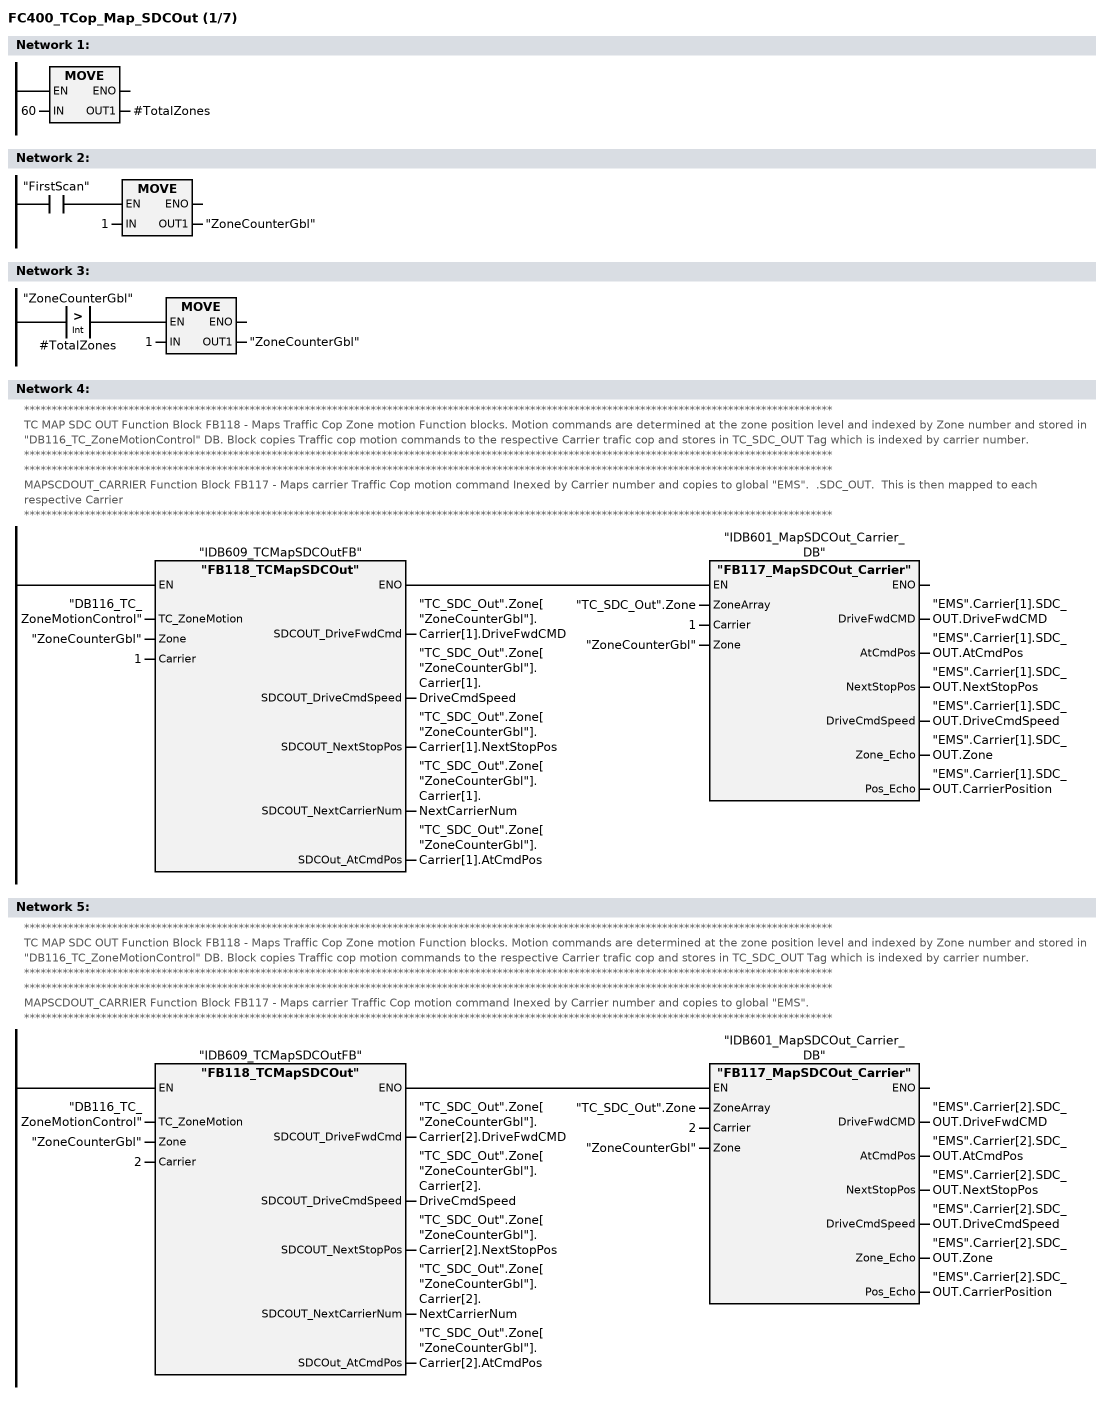
   RUNG wire#powerrail
      Move(in := 60, out1 => #TotalZones)
   END_RUNG
   // the same network as SCL:
   #TotalZones := 60;
END_REGION

REGION Network 2
   RUNG wire#powerrail
      Contact( "FirstScan" )
      Move(in := 1, out1 => "ZoneCounterGbl")
   END_RUNG
   // the same network as SCL:
   IF "FirstScan" THEN "ZoneCounterGbl" := 1; END_IF;
END_REGION

REGION Network 3
   RUNG wire#powerrail
      { S7_Templates := "SrcType := Int" } GT_Contact(in1 := "ZoneCounterGbl", in2 := #TotalZones)
      Move(in := 1, out1 => "ZoneCounterGbl")
   END_RUNG
   // the same network as SCL:
   IF "ZoneCounterGbl" > #TotalZones THEN "ZoneCounterGbl" := 1; END_IF;
END_REGION

REGION Network 4
   // ***************************************************************************************************************************************************
   // 
   // TC MAP SDC OUT Function Block FB118 - Maps Traffic Cop Zone motion Function blocks. Motion commands are determined at the zone position level and indexed by Zone number and stored in 
   //  "DB116_TC_ZoneMotionControl" DB. Block copies Traffic cop motion commands to the respective Carrier trafic cop and stores in TC_SDC_OUT Tag which is indexed by carrier number. 
   // 
   // ***************************************************************************************************************************************************
   // 
   // ***************************************************************************************************************************************************
   // 
   // MAPSCDOUT_CARRIER Function Block FB117 - Maps carrier Traffic Cop motion command Inexed by Carrier number and copies to global "EMS".  .SDC_OUT.  This is then mapped to each respective Carrier
   // 
   // ***************************************************************************************************************************************************
   RUNG wire#powerrail
      "IDB609_TCMapSDCOutFB"(TC_ZoneMotion := "DB116_TC_ZoneMotionControl", Zone := "ZoneCounterGbl", Carrier := 1, SDCOUT_DriveFwdCmd => "TC_SDC_Out".Zone["ZoneCounterGbl"].Carrier[1].DriveFwdCMD, SDCOUT_DriveCmdSpeed => "TC_SDC_Out".Zone["ZoneCounterGbl"].Carrier[1].DriveCmdSpeed, SDCOUT_NextStopPos => "TC_SDC_Out".Zone["ZoneCounterGbl"].Carrier[1].NextStopPos, SDCOUT_NextCarrierNum => "TC_SDC_Out".Zone["ZoneCounterGbl"].Carrier[1].NextCarrierNum, SDCOut_AtCmdPos => "TC_SDC_Out".Zone["ZoneCounterGbl"].Carrier[1].AtCmdPos)
      "IDB601_MapSDCOut_Carrier_DB"(ZoneArray := "TC_SDC_Out".Zone, Carrier := 1, Zone := "ZoneCounterGbl", DriveFwdCMD => "EMS".Carrier[1].SDC_OUT.DriveFwdCMD, AtCmdPos => "EMS".Carrier[1].SDC_OUT.AtCmdPos, NextStopPos => "EMS".Carrier[1].SDC_OUT.NextStopPos, DriveCmdSpeed => "EMS".Carrier[1].SDC_OUT.DriveCmdSpeed, Zone_Echo => "EMS".Carrier[1].SDC_OUT.Zone, Pos_Echo => "EMS".Carrier[1].SDC_OUT.CarrierPosition)
   END_RUNG
   // the same network as SCL:
   "IDB609_TCMapSDCOutFB"(TC_ZoneMotion := "DB116_TC_ZoneMotionControl",   // "FB118_TCMapSDCOut"
                          Zone := "ZoneCounterGbl",
                          Carrier := 1,
                          SDCOUT_DriveFwdCmd => "TC_SDC_Out".Zone["ZoneCounterGbl"].Carrier[1].DriveFwdCMD,
                          SDCOUT_DriveCmdSpeed => "TC_SDC_Out".Zone["ZoneCounterGbl"].Carrier[1].DriveCmdSpeed,
                          SDCOUT_NextStopPos => "TC_SDC_Out".Zone["ZoneCounterGbl"].Carrier[1].NextStopPos,
                          SDCOUT_NextCarrierNum => "TC_SDC_Out".Zone["ZoneCounterGbl"].Carrier[1].NextCarrierNum,
                          SDCOut_AtCmdPos => "TC_SDC_Out".Zone["ZoneCounterGbl"].Carrier[1].AtCmdPos,
                          ENO => #_w1);
   IF #_w1 THEN
       "IDB601_MapSDCOut_Carrier_DB"(ZoneArray := "TC_SDC_Out".Zone,   // "FB117_MapSDCOut_Carrier"
                               Carrier := 1,
                               Zone := "ZoneCounterGbl",
                               DriveFwdCMD => "EMS".Carrier[1].SDC_OUT.DriveFwdCMD,
                               AtCmdPos => "EMS".Carrier[1].SDC_OUT.AtCmdPos,
                               NextStopPos => "EMS".Carrier[1].SDC_OUT.NextStopPos,
                               DriveCmdSpeed => "EMS".Carrier[1].SDC_OUT.DriveCmdSpeed,
                               Zone_Echo => "EMS".Carrier[1].SDC_OUT.Zone,
                               Pos_Echo => "EMS".Carrier[1].SDC_OUT.CarrierPosition);
   END_IF;
END_REGION

REGION Network 5
   // ***************************************************************************************************************************************************
   // 
   // TC MAP SDC OUT Function Block FB118 - Maps Traffic Cop Zone motion Function blocks. Motion commands are determined at the zone position level and indexed by Zone number and stored in 
   //  "DB116_TC_ZoneMotionControl" DB. Block copies Traffic cop motion commands to the respective Carrier trafic cop and stores in TC_SDC_OUT Tag which is indexed by carrier number. 
   // 
   // ***************************************************************************************************************************************************
   // 
   // ***************************************************************************************************************************************************
   // 
   // MAPSCDOUT_CARRIER Function Block FB117 - Maps carrier Traffic Cop motion command Inexed by Carrier number and copies to global "EMS". 
   // 
   // ***************************************************************************************************************************************************
   RUNG wire#powerrail
      "IDB609_TCMapSDCOutFB"(TC_ZoneMotion := "DB116_TC_ZoneMotionControl", Zone := "ZoneCounterGbl", Carrier := 2, SDCOUT_DriveFwdCmd => "TC_SDC_Out".Zone["ZoneCounterGbl"].Carrier[2].DriveFwdCMD, SDCOUT_DriveCmdSpeed => "TC_SDC_Out".Zone["ZoneCounterGbl"].Carrier[2].DriveCmdSpeed, SDCOUT_NextStopPos => "TC_SDC_Out".Zone["ZoneCounterGbl"].Carrier[2].NextStopPos, SDCOUT_NextCarrierNum => "TC_SDC_Out".Zone["ZoneCounterGbl"].Carrier[2].NextCarrierNum, SDCOut_AtCmdPos => "TC_SDC_Out".Zone["ZoneCounterGbl"].Carrier[2].AtCmdPos)
      "IDB601_MapSDCOut_Carrier_DB"(ZoneArray := "TC_SDC_Out".Zone, Carrier := 2, Zone := "ZoneCounterGbl", DriveFwdCMD => "EMS".Carrier[2].SDC_OUT.DriveFwdCMD, AtCmdPos => "EMS".Carrier[2].SDC_OUT.AtCmdPos, NextStopPos => "EMS".Carrier[2].SDC_OUT.NextStopPos, DriveCmdSpeed => "EMS".Carrier[2].SDC_OUT.DriveCmdSpeed, Zone_Echo => "EMS".Carrier[2].SDC_OUT.Zone, Pos_Echo => "EMS".Carrier[2].SDC_OUT.CarrierPosition)
   END_RUNG
   // the same network as SCL:
   "IDB609_TCMapSDCOutFB"(TC_ZoneMotion := "DB116_TC_ZoneMotionControl",   // "FB118_TCMapSDCOut"
                          Zone := "ZoneCounterGbl",
                          Carrier := 2,
                          SDCOUT_DriveFwdCmd => "TC_SDC_Out".Zone["ZoneCounterGbl"].Carrier[2].DriveFwdCMD,
                          SDCOUT_DriveCmdSpeed => "TC_SDC_Out".Zone["ZoneCounterGbl"].Carrier[2].DriveCmdSpeed,
                          SDCOUT_NextStopPos => "TC_SDC_Out".Zone["ZoneCounterGbl"].Carrier[2].NextStopPos,
                          SDCOUT_NextCarrierNum => "TC_SDC_Out".Zone["ZoneCounterGbl"].Carrier[2].NextCarrierNum,
                          SDCOut_AtCmdPos => "TC_SDC_Out".Zone["ZoneCounterGbl"].Carrier[2].AtCmdPos,
                          ENO => #_w1);
   IF #_w1 THEN
       "IDB601_MapSDCOut_Carrier_DB"(ZoneArray := "TC_SDC_Out".Zone,   // "FB117_MapSDCOut_Carrier"
                               Carrier := 2,
                               Zone := "ZoneCounterGbl",
                               DriveFwdCMD => "EMS".Carrier[2].SDC_OUT.DriveFwdCMD,
                               AtCmdPos => "EMS".Carrier[2].SDC_OUT.AtCmdPos,
                               NextStopPos => "EMS".Carrier[2].SDC_OUT.NextStopPos,
                               DriveCmdSpeed => "EMS".Carrier[2].SDC_OUT.DriveCmdSpeed,
                               Zone_Echo => "EMS".Carrier[2].SDC_OUT.Zone,
                               Pos_Echo => "EMS".Carrier[2].SDC_OUT.CarrierPosition);
   END_IF;
END_REGION

REGION Network 6
   // ***************************************************************************************************************************************************
   // 
   // TC MAP SDC OUT Function Block FB118 - Maps Traffic Cop Zone motion Function blocks. Motion commands are determined at the zone position level and indexed by Zone number and stored in 
   //  "DB116_TC_ZoneMotionControl" DB. Block copies Traffic cop motion commands to the respective Carrier trafic cop and stores in TC_SDC_OUT Tag which is indexed by carrier number. 
   // 
   // ***************************************************************************************************************************************************
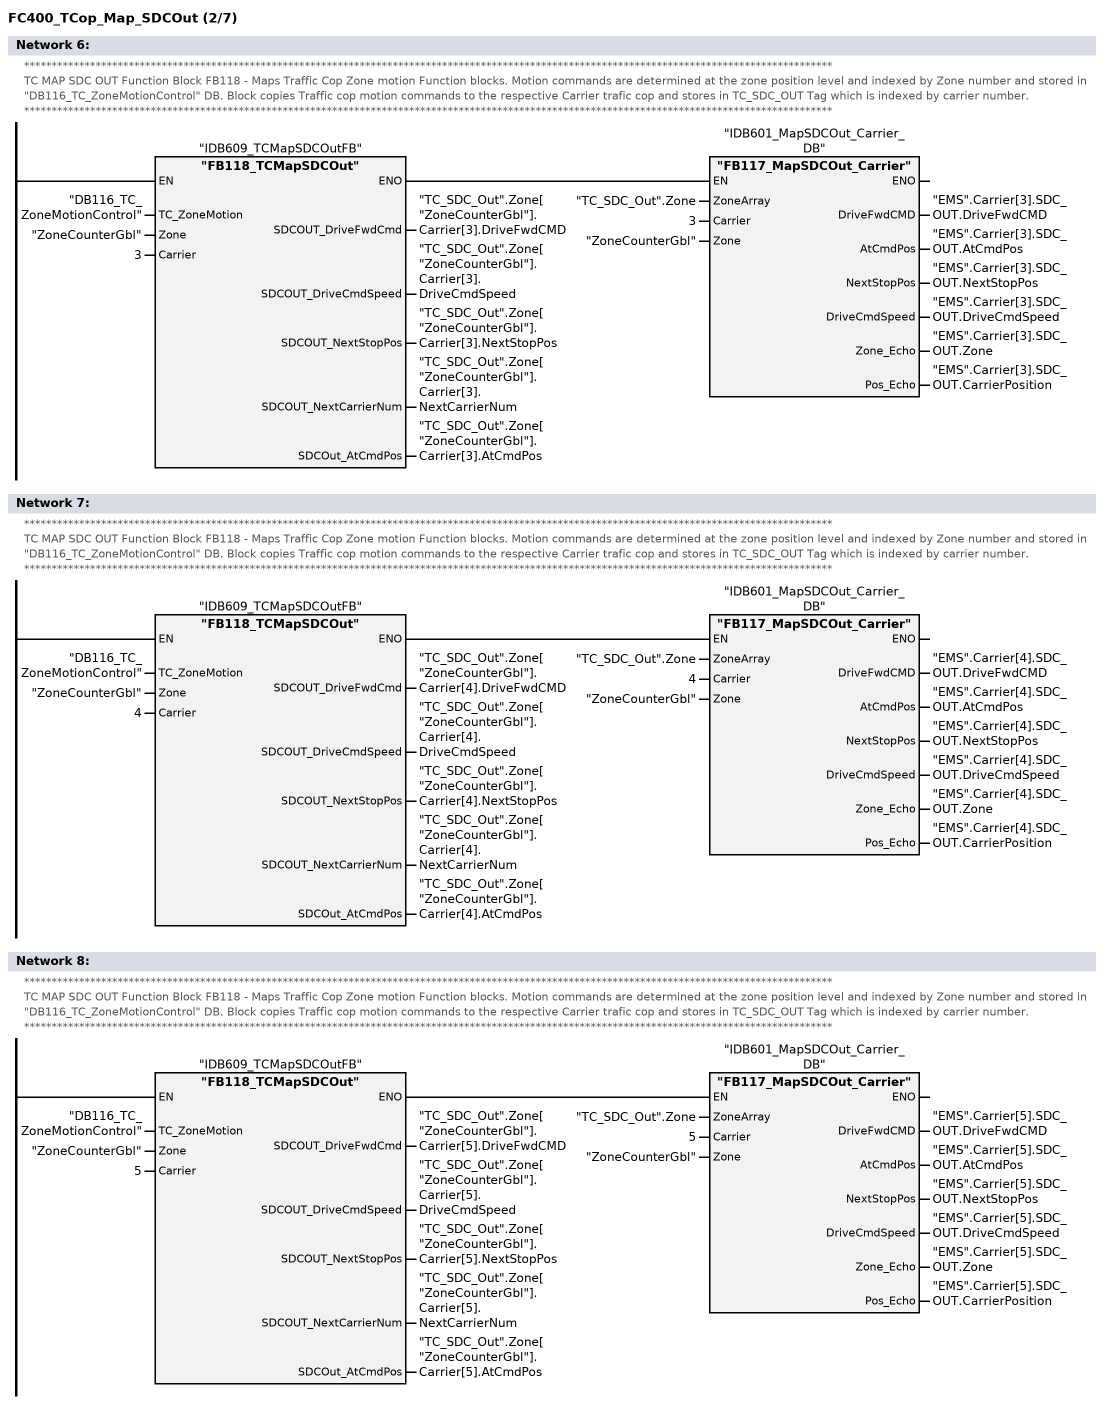
   RUNG wire#powerrail
      "IDB609_TCMapSDCOutFB"(TC_ZoneMotion := "DB116_TC_ZoneMotionControl", Zone := "ZoneCounterGbl", Carrier := 3, SDCOUT_DriveFwdCmd => "TC_SDC_Out".Zone["ZoneCounterGbl"].Carrier[3].DriveFwdCMD, SDCOUT_DriveCmdSpeed => "TC_SDC_Out".Zone["ZoneCounterGbl"].Carrier[3].DriveCmdSpeed, SDCOUT_NextStopPos => "TC_SDC_Out".Zone["ZoneCounterGbl"].Carrier[3].NextStopPos, SDCOUT_NextCarrierNum => "TC_SDC_Out".Zone["ZoneCounterGbl"].Carrier[3].NextCarrierNum, SDCOut_AtCmdPos => "TC_SDC_Out".Zone["ZoneCounterGbl"].Carrier[3].AtCmdPos)
      "IDB601_MapSDCOut_Carrier_DB"(ZoneArray := "TC_SDC_Out".Zone, Carrier := 3, Zone := "ZoneCounterGbl", DriveFwdCMD => "EMS".Carrier[3].SDC_OUT.DriveFwdCMD, AtCmdPos => "EMS".Carrier[3].SDC_OUT.AtCmdPos, NextStopPos => "EMS".Carrier[3].SDC_OUT.NextStopPos, DriveCmdSpeed => "EMS".Carrier[3].SDC_OUT.DriveCmdSpeed, Zone_Echo => "EMS".Carrier[3].SDC_OUT.Zone, Pos_Echo => "EMS".Carrier[3].SDC_OUT.CarrierPosition)
   END_RUNG
   // the same network as SCL:
   "IDB609_TCMapSDCOutFB"(TC_ZoneMotion := "DB116_TC_ZoneMotionControl",   // "FB118_TCMapSDCOut"
                          Zone := "ZoneCounterGbl",
                          Carrier := 3,
                          SDCOUT_DriveFwdCmd => "TC_SDC_Out".Zone["ZoneCounterGbl"].Carrier[3].DriveFwdCMD,
                          SDCOUT_DriveCmdSpeed => "TC_SDC_Out".Zone["ZoneCounterGbl"].Carrier[3].DriveCmdSpeed,
                          SDCOUT_NextStopPos => "TC_SDC_Out".Zone["ZoneCounterGbl"].Carrier[3].NextStopPos,
                          SDCOUT_NextCarrierNum => "TC_SDC_Out".Zone["ZoneCounterGbl"].Carrier[3].NextCarrierNum,
                          SDCOut_AtCmdPos => "TC_SDC_Out".Zone["ZoneCounterGbl"].Carrier[3].AtCmdPos,
                          ENO => #_w1);
   IF #_w1 THEN
       "IDB601_MapSDCOut_Carrier_DB"(ZoneArray := "TC_SDC_Out".Zone,   // "FB117_MapSDCOut_Carrier"
                               Carrier := 3,
                               Zone := "ZoneCounterGbl",
                               DriveFwdCMD => "EMS".Carrier[3].SDC_OUT.DriveFwdCMD,
                               AtCmdPos => "EMS".Carrier[3].SDC_OUT.AtCmdPos,
                               NextStopPos => "EMS".Carrier[3].SDC_OUT.NextStopPos,
                               DriveCmdSpeed => "EMS".Carrier[3].SDC_OUT.DriveCmdSpeed,
                               Zone_Echo => "EMS".Carrier[3].SDC_OUT.Zone,
                               Pos_Echo => "EMS".Carrier[3].SDC_OUT.CarrierPosition);
   END_IF;
END_REGION

REGION Network 7
   // ***************************************************************************************************************************************************
   // 
   // TC MAP SDC OUT Function Block FB118 - Maps Traffic Cop Zone motion Function blocks. Motion commands are determined at the zone position level and indexed by Zone number and stored in 
   //  "DB116_TC_ZoneMotionControl" DB. Block copies Traffic cop motion commands to the respective Carrier trafic cop and stores in TC_SDC_OUT Tag which is indexed by carrier number. 
   // 
   // ***************************************************************************************************************************************************
   RUNG wire#powerrail
      "IDB609_TCMapSDCOutFB"(TC_ZoneMotion := "DB116_TC_ZoneMotionControl", Zone := "ZoneCounterGbl", Carrier := 4, SDCOUT_DriveFwdCmd => "TC_SDC_Out".Zone["ZoneCounterGbl"].Carrier[4].DriveFwdCMD, SDCOUT_DriveCmdSpeed => "TC_SDC_Out".Zone["ZoneCounterGbl"].Carrier[4].DriveCmdSpeed, SDCOUT_NextStopPos => "TC_SDC_Out".Zone["ZoneCounterGbl"].Carrier[4].NextStopPos, SDCOUT_NextCarrierNum => "TC_SDC_Out".Zone["ZoneCounterGbl"].Carrier[4].NextCarrierNum, SDCOut_AtCmdPos => "TC_SDC_Out".Zone["ZoneCounterGbl"].Carrier[4].AtCmdPos)
      "IDB601_MapSDCOut_Carrier_DB"(ZoneArray := "TC_SDC_Out".Zone, Carrier := 4, Zone := "ZoneCounterGbl", DriveFwdCMD => "EMS".Carrier[4].SDC_OUT.DriveFwdCMD, AtCmdPos => "EMS".Carrier[4].SDC_OUT.AtCmdPos, NextStopPos => "EMS".Carrier[4].SDC_OUT.NextStopPos, DriveCmdSpeed => "EMS".Carrier[4].SDC_OUT.DriveCmdSpeed, Zone_Echo => "EMS".Carrier[4].SDC_OUT.Zone, Pos_Echo => "EMS".Carrier[4].SDC_OUT.CarrierPosition)
   END_RUNG
   // the same network as SCL:
   "IDB609_TCMapSDCOutFB"(TC_ZoneMotion := "DB116_TC_ZoneMotionControl",   // "FB118_TCMapSDCOut"
                          Zone := "ZoneCounterGbl",
                          Carrier := 4,
                          SDCOUT_DriveFwdCmd => "TC_SDC_Out".Zone["ZoneCounterGbl"].Carrier[4].DriveFwdCMD,
                          SDCOUT_DriveCmdSpeed => "TC_SDC_Out".Zone["ZoneCounterGbl"].Carrier[4].DriveCmdSpeed,
                          SDCOUT_NextStopPos => "TC_SDC_Out".Zone["ZoneCounterGbl"].Carrier[4].NextStopPos,
                          SDCOUT_NextCarrierNum => "TC_SDC_Out".Zone["ZoneCounterGbl"].Carrier[4].NextCarrierNum,
                          SDCOut_AtCmdPos => "TC_SDC_Out".Zone["ZoneCounterGbl"].Carrier[4].AtCmdPos,
                          ENO => #_w1);
   IF #_w1 THEN
       "IDB601_MapSDCOut_Carrier_DB"(ZoneArray := "TC_SDC_Out".Zone,   // "FB117_MapSDCOut_Carrier"
                               Carrier := 4,
                               Zone := "ZoneCounterGbl",
                               DriveFwdCMD => "EMS".Carrier[4].SDC_OUT.DriveFwdCMD,
                               AtCmdPos => "EMS".Carrier[4].SDC_OUT.AtCmdPos,
                               NextStopPos => "EMS".Carrier[4].SDC_OUT.NextStopPos,
                               DriveCmdSpeed => "EMS".Carrier[4].SDC_OUT.DriveCmdSpeed,
                               Zone_Echo => "EMS".Carrier[4].SDC_OUT.Zone,
                               Pos_Echo => "EMS".Carrier[4].SDC_OUT.CarrierPosition);
   END_IF;
END_REGION

REGION Network 8
   // ***************************************************************************************************************************************************
   // 
   // TC MAP SDC OUT Function Block FB118 - Maps Traffic Cop Zone motion Function blocks. Motion commands are determined at the zone position level and indexed by Zone number and stored in 
   //  "DB116_TC_ZoneMotionControl" DB. Block copies Traffic cop motion commands to the respective Carrier trafic cop and stores in TC_SDC_OUT Tag which is indexed by carrier number. 
   // 
   // ***************************************************************************************************************************************************
   RUNG wire#powerrail
      "IDB609_TCMapSDCOutFB"(TC_ZoneMotion := "DB116_TC_ZoneMotionControl", Zone := "ZoneCounterGbl", Carrier := 5, SDCOUT_DriveFwdCmd => "TC_SDC_Out".Zone["ZoneCounterGbl"].Carrier[5].DriveFwdCMD, SDCOUT_DriveCmdSpeed => "TC_SDC_Out".Zone["ZoneCounterGbl"].Carrier[5].DriveCmdSpeed, SDCOUT_NextStopPos => "TC_SDC_Out".Zone["ZoneCounterGbl"].Carrier[5].NextStopPos, SDCOUT_NextCarrierNum => "TC_SDC_Out".Zone["ZoneCounterGbl"].Carrier[5].NextCarrierNum, SDCOut_AtCmdPos => "TC_SDC_Out".Zone["ZoneCounterGbl"].Carrier[5].AtCmdPos)
      "IDB601_MapSDCOut_Carrier_DB"(ZoneArray := "TC_SDC_Out".Zone, Carrier := 5, Zone := "ZoneCounterGbl", DriveFwdCMD => "EMS".Carrier[5].SDC_OUT.DriveFwdCMD, AtCmdPos => "EMS".Carrier[5].SDC_OUT.AtCmdPos, NextStopPos => "EMS".Carrier[5].SDC_OUT.NextStopPos, DriveCmdSpeed => "EMS".Carrier[5].SDC_OUT.DriveCmdSpeed, Zone_Echo => "EMS".Carrier[5].SDC_OUT.Zone, Pos_Echo => "EMS".Carrier[5].SDC_OUT.CarrierPosition)
   END_RUNG
   // the same network as SCL:
   "IDB609_TCMapSDCOutFB"(TC_ZoneMotion := "DB116_TC_ZoneMotionControl",   // "FB118_TCMapSDCOut"
                          Zone := "ZoneCounterGbl",
                          Carrier := 5,
                          SDCOUT_DriveFwdCmd => "TC_SDC_Out".Zone["ZoneCounterGbl"].Carrier[5].DriveFwdCMD,
                          SDCOUT_DriveCmdSpeed => "TC_SDC_Out".Zone["ZoneCounterGbl"].Carrier[5].DriveCmdSpeed,
                          SDCOUT_NextStopPos => "TC_SDC_Out".Zone["ZoneCounterGbl"].Carrier[5].NextStopPos,
                          SDCOUT_NextCarrierNum => "TC_SDC_Out".Zone["ZoneCounterGbl"].Carrier[5].NextCarrierNum,
                          SDCOut_AtCmdPos => "TC_SDC_Out".Zone["ZoneCounterGbl"].Carrier[5].AtCmdPos,
                          ENO => #_w1);
   IF #_w1 THEN
       "IDB601_MapSDCOut_Carrier_DB"(ZoneArray := "TC_SDC_Out".Zone,   // "FB117_MapSDCOut_Carrier"
                               Carrier := 5,
                               Zone := "ZoneCounterGbl",
                               DriveFwdCMD => "EMS".Carrier[5].SDC_OUT.DriveFwdCMD,
                               AtCmdPos => "EMS".Carrier[5].SDC_OUT.AtCmdPos,
                               NextStopPos => "EMS".Carrier[5].SDC_OUT.NextStopPos,
                               DriveCmdSpeed => "EMS".Carrier[5].SDC_OUT.DriveCmdSpeed,
                               Zone_Echo => "EMS".Carrier[5].SDC_OUT.Zone,
                               Pos_Echo => "EMS".Carrier[5].SDC_OUT.CarrierPosition);
   END_IF;
END_REGION

REGION Network 9
   // ***************************************************************************************************************************************************
   // 
   // TC MAP SDC OUT Function Block FB118 - Maps Traffic Cop Zone motion Function blocks. Motion commands are determined at the zone position level and indexed by Zone number and stored in 
   //  "DB116_TC_ZoneMotionControl" DB. Block copies Traffic cop motion commands to the respective Carrier trafic cop and stores in TC_SDC_OUT Tag which is indexed by carrier number. 
   // 
   // ***************************************************************************************************************************************************
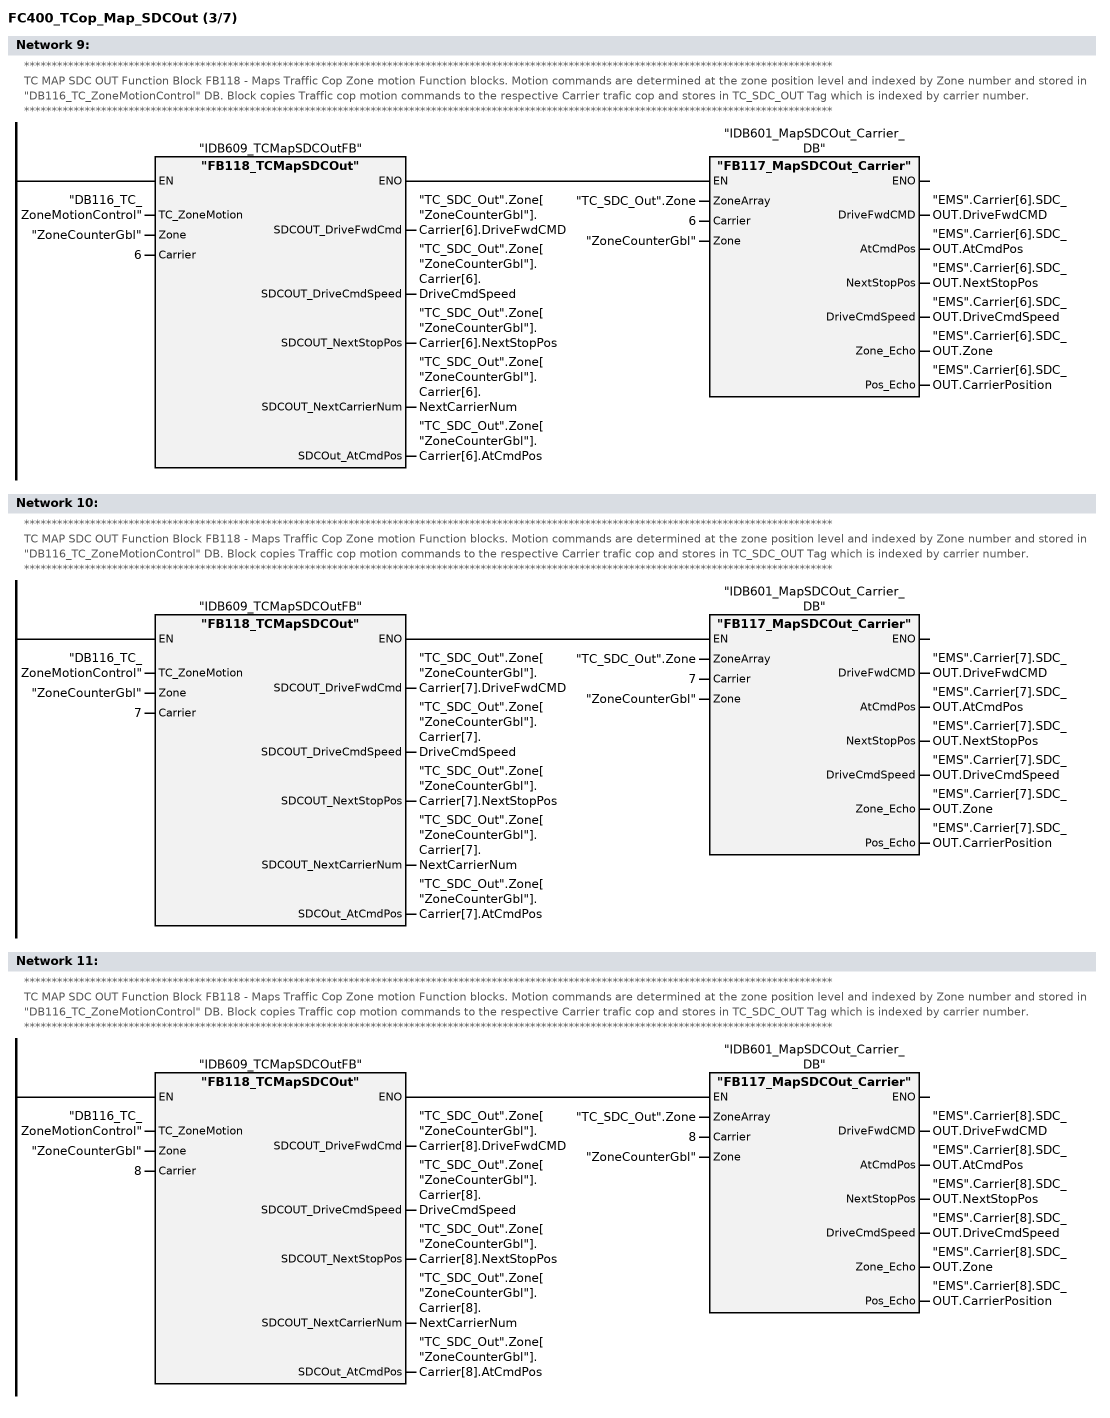
   RUNG wire#powerrail
      "IDB609_TCMapSDCOutFB"(TC_ZoneMotion := "DB116_TC_ZoneMotionControl", Zone := "ZoneCounterGbl", Carrier := 6, SDCOUT_DriveFwdCmd => "TC_SDC_Out".Zone["ZoneCounterGbl"].Carrier[6].DriveFwdCMD, SDCOUT_DriveCmdSpeed => "TC_SDC_Out".Zone["ZoneCounterGbl"].Carrier[6].DriveCmdSpeed, SDCOUT_NextStopPos => "TC_SDC_Out".Zone["ZoneCounterGbl"].Carrier[6].NextStopPos, SDCOUT_NextCarrierNum => "TC_SDC_Out".Zone["ZoneCounterGbl"].Carrier[6].NextCarrierNum, SDCOut_AtCmdPos => "TC_SDC_Out".Zone["ZoneCounterGbl"].Carrier[6].AtCmdPos)
      "IDB601_MapSDCOut_Carrier_DB"(ZoneArray := "TC_SDC_Out".Zone, Carrier := 6, Zone := "ZoneCounterGbl", DriveFwdCMD => "EMS".Carrier[6].SDC_OUT.DriveFwdCMD, AtCmdPos => "EMS".Carrier[6].SDC_OUT.AtCmdPos, NextStopPos => "EMS".Carrier[6].SDC_OUT.NextStopPos, DriveCmdSpeed => "EMS".Carrier[6].SDC_OUT.DriveCmdSpeed, Zone_Echo => "EMS".Carrier[6].SDC_OUT.Zone, Pos_Echo => "EMS".Carrier[6].SDC_OUT.CarrierPosition)
   END_RUNG
   // the same network as SCL:
   "IDB609_TCMapSDCOutFB"(TC_ZoneMotion := "DB116_TC_ZoneMotionControl",   // "FB118_TCMapSDCOut"
                          Zone := "ZoneCounterGbl",
                          Carrier := 6,
                          SDCOUT_DriveFwdCmd => "TC_SDC_Out".Zone["ZoneCounterGbl"].Carrier[6].DriveFwdCMD,
                          SDCOUT_DriveCmdSpeed => "TC_SDC_Out".Zone["ZoneCounterGbl"].Carrier[6].DriveCmdSpeed,
                          SDCOUT_NextStopPos => "TC_SDC_Out".Zone["ZoneCounterGbl"].Carrier[6].NextStopPos,
                          SDCOUT_NextCarrierNum => "TC_SDC_Out".Zone["ZoneCounterGbl"].Carrier[6].NextCarrierNum,
                          SDCOut_AtCmdPos => "TC_SDC_Out".Zone["ZoneCounterGbl"].Carrier[6].AtCmdPos,
                          ENO => #_w1);
   IF #_w1 THEN
       "IDB601_MapSDCOut_Carrier_DB"(ZoneArray := "TC_SDC_Out".Zone,   // "FB117_MapSDCOut_Carrier"
                               Carrier := 6,
                               Zone := "ZoneCounterGbl",
                               DriveFwdCMD => "EMS".Carrier[6].SDC_OUT.DriveFwdCMD,
                               AtCmdPos => "EMS".Carrier[6].SDC_OUT.AtCmdPos,
                               NextStopPos => "EMS".Carrier[6].SDC_OUT.NextStopPos,
                               DriveCmdSpeed => "EMS".Carrier[6].SDC_OUT.DriveCmdSpeed,
                               Zone_Echo => "EMS".Carrier[6].SDC_OUT.Zone,
                               Pos_Echo => "EMS".Carrier[6].SDC_OUT.CarrierPosition);
   END_IF;
END_REGION

REGION Network 10
   // ***************************************************************************************************************************************************
   // 
   // TC MAP SDC OUT Function Block FB118 - Maps Traffic Cop Zone motion Function blocks. Motion commands are determined at the zone position level and indexed by Zone number and stored in 
   //  "DB116_TC_ZoneMotionControl" DB. Block copies Traffic cop motion commands to the respective Carrier trafic cop and stores in TC_SDC_OUT Tag which is indexed by carrier number. 
   // 
   // ***************************************************************************************************************************************************
   RUNG wire#powerrail
      "IDB609_TCMapSDCOutFB"(TC_ZoneMotion := "DB116_TC_ZoneMotionControl", Zone := "ZoneCounterGbl", Carrier := 7, SDCOUT_DriveFwdCmd => "TC_SDC_Out".Zone["ZoneCounterGbl"].Carrier[7].DriveFwdCMD, SDCOUT_DriveCmdSpeed => "TC_SDC_Out".Zone["ZoneCounterGbl"].Carrier[7].DriveCmdSpeed, SDCOUT_NextStopPos => "TC_SDC_Out".Zone["ZoneCounterGbl"].Carrier[7].NextStopPos, SDCOUT_NextCarrierNum => "TC_SDC_Out".Zone["ZoneCounterGbl"].Carrier[7].NextCarrierNum, SDCOut_AtCmdPos => "TC_SDC_Out".Zone["ZoneCounterGbl"].Carrier[7].AtCmdPos)
      "IDB601_MapSDCOut_Carrier_DB"(ZoneArray := "TC_SDC_Out".Zone, Carrier := 7, Zone := "ZoneCounterGbl", DriveFwdCMD => "EMS".Carrier[7].SDC_OUT.DriveFwdCMD, AtCmdPos => "EMS".Carrier[7].SDC_OUT.AtCmdPos, NextStopPos => "EMS".Carrier[7].SDC_OUT.NextStopPos, DriveCmdSpeed => "EMS".Carrier[7].SDC_OUT.DriveCmdSpeed, Zone_Echo => "EMS".Carrier[7].SDC_OUT.Zone, Pos_Echo => "EMS".Carrier[7].SDC_OUT.CarrierPosition)
   END_RUNG
   // the same network as SCL:
   "IDB609_TCMapSDCOutFB"(TC_ZoneMotion := "DB116_TC_ZoneMotionControl",   // "FB118_TCMapSDCOut"
                          Zone := "ZoneCounterGbl",
                          Carrier := 7,
                          SDCOUT_DriveFwdCmd => "TC_SDC_Out".Zone["ZoneCounterGbl"].Carrier[7].DriveFwdCMD,
                          SDCOUT_DriveCmdSpeed => "TC_SDC_Out".Zone["ZoneCounterGbl"].Carrier[7].DriveCmdSpeed,
                          SDCOUT_NextStopPos => "TC_SDC_Out".Zone["ZoneCounterGbl"].Carrier[7].NextStopPos,
                          SDCOUT_NextCarrierNum => "TC_SDC_Out".Zone["ZoneCounterGbl"].Carrier[7].NextCarrierNum,
                          SDCOut_AtCmdPos => "TC_SDC_Out".Zone["ZoneCounterGbl"].Carrier[7].AtCmdPos,
                          ENO => #_w1);
   IF #_w1 THEN
       "IDB601_MapSDCOut_Carrier_DB"(ZoneArray := "TC_SDC_Out".Zone,   // "FB117_MapSDCOut_Carrier"
                               Carrier := 7,
                               Zone := "ZoneCounterGbl",
                               DriveFwdCMD => "EMS".Carrier[7].SDC_OUT.DriveFwdCMD,
                               AtCmdPos => "EMS".Carrier[7].SDC_OUT.AtCmdPos,
                               NextStopPos => "EMS".Carrier[7].SDC_OUT.NextStopPos,
                               DriveCmdSpeed => "EMS".Carrier[7].SDC_OUT.DriveCmdSpeed,
                               Zone_Echo => "EMS".Carrier[7].SDC_OUT.Zone,
                               Pos_Echo => "EMS".Carrier[7].SDC_OUT.CarrierPosition);
   END_IF;
END_REGION

REGION Network 11
   // ***************************************************************************************************************************************************
   // 
   // TC MAP SDC OUT Function Block FB118 - Maps Traffic Cop Zone motion Function blocks. Motion commands are determined at the zone position level and indexed by Zone number and stored in 
   //  "DB116_TC_ZoneMotionControl" DB. Block copies Traffic cop motion commands to the respective Carrier trafic cop and stores in TC_SDC_OUT Tag which is indexed by carrier number. 
   // 
   // ***************************************************************************************************************************************************
   RUNG wire#powerrail
      "IDB609_TCMapSDCOutFB"(TC_ZoneMotion := "DB116_TC_ZoneMotionControl", Zone := "ZoneCounterGbl", Carrier := 8, SDCOUT_DriveFwdCmd => "TC_SDC_Out".Zone["ZoneCounterGbl"].Carrier[8].DriveFwdCMD, SDCOUT_DriveCmdSpeed => "TC_SDC_Out".Zone["ZoneCounterGbl"].Carrier[8].DriveCmdSpeed, SDCOUT_NextStopPos => "TC_SDC_Out".Zone["ZoneCounterGbl"].Carrier[8].NextStopPos, SDCOUT_NextCarrierNum => "TC_SDC_Out".Zone["ZoneCounterGbl"].Carrier[8].NextCarrierNum, SDCOut_AtCmdPos => "TC_SDC_Out".Zone["ZoneCounterGbl"].Carrier[8].AtCmdPos)
      "IDB601_MapSDCOut_Carrier_DB"(ZoneArray := "TC_SDC_Out".Zone, Carrier := 8, Zone := "ZoneCounterGbl", DriveFwdCMD => "EMS".Carrier[8].SDC_OUT.DriveFwdCMD, AtCmdPos => "EMS".Carrier[8].SDC_OUT.AtCmdPos, NextStopPos => "EMS".Carrier[8].SDC_OUT.NextStopPos, DriveCmdSpeed => "EMS".Carrier[8].SDC_OUT.DriveCmdSpeed, Zone_Echo => "EMS".Carrier[8].SDC_OUT.Zone, Pos_Echo => "EMS".Carrier[8].SDC_OUT.CarrierPosition)
   END_RUNG
   // the same network as SCL:
   "IDB609_TCMapSDCOutFB"(TC_ZoneMotion := "DB116_TC_ZoneMotionControl",   // "FB118_TCMapSDCOut"
                          Zone := "ZoneCounterGbl",
                          Carrier := 8,
                          SDCOUT_DriveFwdCmd => "TC_SDC_Out".Zone["ZoneCounterGbl"].Carrier[8].DriveFwdCMD,
                          SDCOUT_DriveCmdSpeed => "TC_SDC_Out".Zone["ZoneCounterGbl"].Carrier[8].DriveCmdSpeed,
                          SDCOUT_NextStopPos => "TC_SDC_Out".Zone["ZoneCounterGbl"].Carrier[8].NextStopPos,
                          SDCOUT_NextCarrierNum => "TC_SDC_Out".Zone["ZoneCounterGbl"].Carrier[8].NextCarrierNum,
                          SDCOut_AtCmdPos => "TC_SDC_Out".Zone["ZoneCounterGbl"].Carrier[8].AtCmdPos,
                          ENO => #_w1);
   IF #_w1 THEN
       "IDB601_MapSDCOut_Carrier_DB"(ZoneArray := "TC_SDC_Out".Zone,   // "FB117_MapSDCOut_Carrier"
                               Carrier := 8,
                               Zone := "ZoneCounterGbl",
                               DriveFwdCMD => "EMS".Carrier[8].SDC_OUT.DriveFwdCMD,
                               AtCmdPos => "EMS".Carrier[8].SDC_OUT.AtCmdPos,
                               NextStopPos => "EMS".Carrier[8].SDC_OUT.NextStopPos,
                               DriveCmdSpeed => "EMS".Carrier[8].SDC_OUT.DriveCmdSpeed,
                               Zone_Echo => "EMS".Carrier[8].SDC_OUT.Zone,
                               Pos_Echo => "EMS".Carrier[8].SDC_OUT.CarrierPosition);
   END_IF;
END_REGION

REGION Network 12
   // ***************************************************************************************************************************************************
   // 
   // TC MAP SDC OUT Function Block FB118 - Maps Traffic Cop Zone motion Function blocks. Motion commands are determined at the zone position level and indexed by Zone number and stored in 
   //  "DB116_TC_ZoneMotionControl" DB. Block copies Traffic cop motion commands to the respective Carrier trafic cop and stores in TC_SDC_OUT Tag which is indexed by carrier number. 
   // 
   // ***************************************************************************************************************************************************
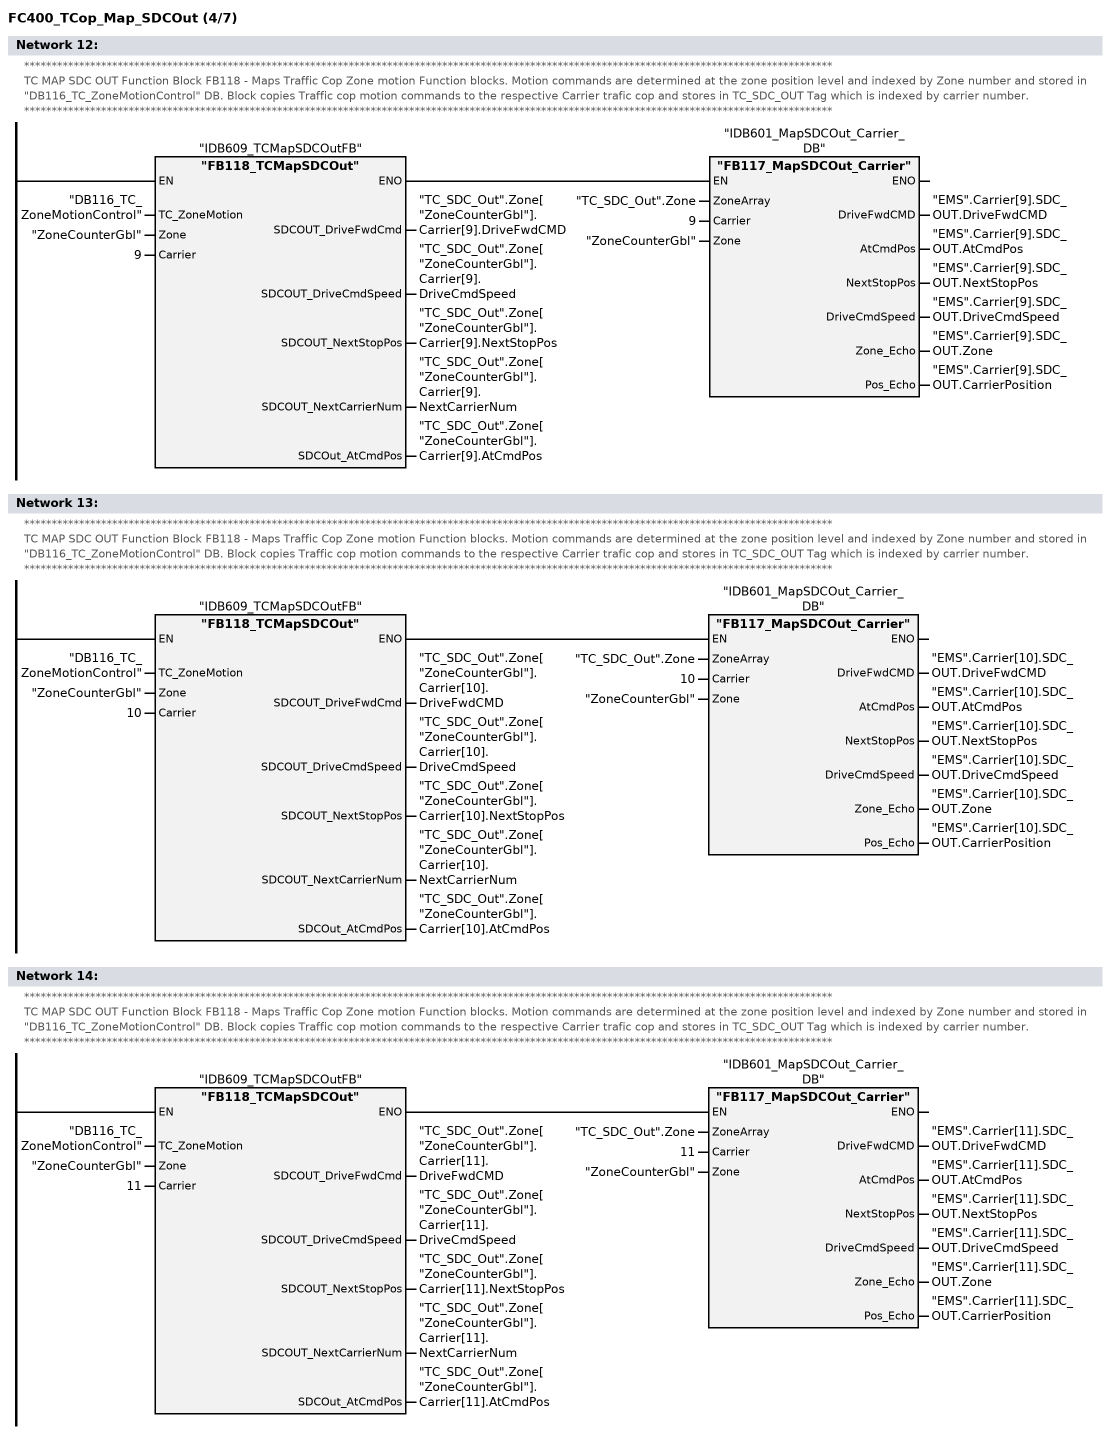
   RUNG wire#powerrail
      "IDB609_TCMapSDCOutFB"(TC_ZoneMotion := "DB116_TC_ZoneMotionControl", Zone := "ZoneCounterGbl", Carrier := 9, SDCOUT_DriveFwdCmd => "TC_SDC_Out".Zone["ZoneCounterGbl"].Carrier[9].DriveFwdCMD, SDCOUT_DriveCmdSpeed => "TC_SDC_Out".Zone["ZoneCounterGbl"].Carrier[9].DriveCmdSpeed, SDCOUT_NextStopPos => "TC_SDC_Out".Zone["ZoneCounterGbl"].Carrier[9].NextStopPos, SDCOUT_NextCarrierNum => "TC_SDC_Out".Zone["ZoneCounterGbl"].Carrier[9].NextCarrierNum, SDCOut_AtCmdPos => "TC_SDC_Out".Zone["ZoneCounterGbl"].Carrier[9].AtCmdPos)
      "IDB601_MapSDCOut_Carrier_DB"(ZoneArray := "TC_SDC_Out".Zone, Carrier := 9, Zone := "ZoneCounterGbl", DriveFwdCMD => "EMS".Carrier[9].SDC_OUT.DriveFwdCMD, AtCmdPos => "EMS".Carrier[9].SDC_OUT.AtCmdPos, NextStopPos => "EMS".Carrier[9].SDC_OUT.NextStopPos, DriveCmdSpeed => "EMS".Carrier[9].SDC_OUT.DriveCmdSpeed, Zone_Echo => "EMS".Carrier[9].SDC_OUT.Zone, Pos_Echo => "EMS".Carrier[9].SDC_OUT.CarrierPosition)
   END_RUNG
   // the same network as SCL:
   "IDB609_TCMapSDCOutFB"(TC_ZoneMotion := "DB116_TC_ZoneMotionControl",   // "FB118_TCMapSDCOut"
                          Zone := "ZoneCounterGbl",
                          Carrier := 9,
                          SDCOUT_DriveFwdCmd => "TC_SDC_Out".Zone["ZoneCounterGbl"].Carrier[9].DriveFwdCMD,
                          SDCOUT_DriveCmdSpeed => "TC_SDC_Out".Zone["ZoneCounterGbl"].Carrier[9].DriveCmdSpeed,
                          SDCOUT_NextStopPos => "TC_SDC_Out".Zone["ZoneCounterGbl"].Carrier[9].NextStopPos,
                          SDCOUT_NextCarrierNum => "TC_SDC_Out".Zone["ZoneCounterGbl"].Carrier[9].NextCarrierNum,
                          SDCOut_AtCmdPos => "TC_SDC_Out".Zone["ZoneCounterGbl"].Carrier[9].AtCmdPos,
                          ENO => #_w1);
   IF #_w1 THEN
       "IDB601_MapSDCOut_Carrier_DB"(ZoneArray := "TC_SDC_Out".Zone,   // "FB117_MapSDCOut_Carrier"
                               Carrier := 9,
                               Zone := "ZoneCounterGbl",
                               DriveFwdCMD => "EMS".Carrier[9].SDC_OUT.DriveFwdCMD,
                               AtCmdPos => "EMS".Carrier[9].SDC_OUT.AtCmdPos,
                               NextStopPos => "EMS".Carrier[9].SDC_OUT.NextStopPos,
                               DriveCmdSpeed => "EMS".Carrier[9].SDC_OUT.DriveCmdSpeed,
                               Zone_Echo => "EMS".Carrier[9].SDC_OUT.Zone,
                               Pos_Echo => "EMS".Carrier[9].SDC_OUT.CarrierPosition);
   END_IF;
END_REGION

REGION Network 13
   // ***************************************************************************************************************************************************
   // 
   // TC MAP SDC OUT Function Block FB118 - Maps Traffic Cop Zone motion Function blocks. Motion commands are determined at the zone position level and indexed by Zone number and stored in 
   //  "DB116_TC_ZoneMotionControl" DB. Block copies Traffic cop motion commands to the respective Carrier trafic cop and stores in TC_SDC_OUT Tag which is indexed by carrier number. 
   // 
   // ***************************************************************************************************************************************************
   RUNG wire#powerrail
      "IDB609_TCMapSDCOutFB"(TC_ZoneMotion := "DB116_TC_ZoneMotionControl", Zone := "ZoneCounterGbl", Carrier := 10, SDCOUT_DriveFwdCmd => "TC_SDC_Out".Zone["ZoneCounterGbl"].Carrier[10].DriveFwdCMD, SDCOUT_DriveCmdSpeed => "TC_SDC_Out".Zone["ZoneCounterGbl"].Carrier[10].DriveCmdSpeed, SDCOUT_NextStopPos => "TC_SDC_Out".Zone["ZoneCounterGbl"].Carrier[10].NextStopPos, SDCOUT_NextCarrierNum => "TC_SDC_Out".Zone["ZoneCounterGbl"].Carrier[10].NextCarrierNum, SDCOut_AtCmdPos => "TC_SDC_Out".Zone["ZoneCounterGbl"].Carrier[10].AtCmdPos)
      "IDB601_MapSDCOut_Carrier_DB"(ZoneArray := "TC_SDC_Out".Zone, Carrier := 10, Zone := "ZoneCounterGbl", DriveFwdCMD => "EMS".Carrier[10].SDC_OUT.DriveFwdCMD, AtCmdPos => "EMS".Carrier[10].SDC_OUT.AtCmdPos, NextStopPos => "EMS".Carrier[10].SDC_OUT.NextStopPos, DriveCmdSpeed => "EMS".Carrier[10].SDC_OUT.DriveCmdSpeed, Zone_Echo => "EMS".Carrier[10].SDC_OUT.Zone, Pos_Echo => "EMS".Carrier[10].SDC_OUT.CarrierPosition)
   END_RUNG
   // the same network as SCL:
   "IDB609_TCMapSDCOutFB"(TC_ZoneMotion := "DB116_TC_ZoneMotionControl",   // "FB118_TCMapSDCOut"
                          Zone := "ZoneCounterGbl",
                          Carrier := 10,
                          SDCOUT_DriveFwdCmd => "TC_SDC_Out".Zone["ZoneCounterGbl"].Carrier[10].DriveFwdCMD,
                          SDCOUT_DriveCmdSpeed => "TC_SDC_Out".Zone["ZoneCounterGbl"].Carrier[10].DriveCmdSpeed,
                          SDCOUT_NextStopPos => "TC_SDC_Out".Zone["ZoneCounterGbl"].Carrier[10].NextStopPos,
                          SDCOUT_NextCarrierNum => "TC_SDC_Out".Zone["ZoneCounterGbl"].Carrier[10].NextCarrierNum,
                          SDCOut_AtCmdPos => "TC_SDC_Out".Zone["ZoneCounterGbl"].Carrier[10].AtCmdPos,
                          ENO => #_w1);
   IF #_w1 THEN
       "IDB601_MapSDCOut_Carrier_DB"(ZoneArray := "TC_SDC_Out".Zone,   // "FB117_MapSDCOut_Carrier"
                               Carrier := 10,
                               Zone := "ZoneCounterGbl",
                               DriveFwdCMD => "EMS".Carrier[10].SDC_OUT.DriveFwdCMD,
                               AtCmdPos => "EMS".Carrier[10].SDC_OUT.AtCmdPos,
                               NextStopPos => "EMS".Carrier[10].SDC_OUT.NextStopPos,
                               DriveCmdSpeed => "EMS".Carrier[10].SDC_OUT.DriveCmdSpeed,
                               Zone_Echo => "EMS".Carrier[10].SDC_OUT.Zone,
                               Pos_Echo => "EMS".Carrier[10].SDC_OUT.CarrierPosition);
   END_IF;
END_REGION

REGION Network 14
   // ***************************************************************************************************************************************************
   // 
   // TC MAP SDC OUT Function Block FB118 - Maps Traffic Cop Zone motion Function blocks. Motion commands are determined at the zone position level and indexed by Zone number and stored in 
   //  "DB116_TC_ZoneMotionControl" DB. Block copies Traffic cop motion commands to the respective Carrier trafic cop and stores in TC_SDC_OUT Tag which is indexed by carrier number. 
   // 
   // ***************************************************************************************************************************************************
   RUNG wire#powerrail
      "IDB609_TCMapSDCOutFB"(TC_ZoneMotion := "DB116_TC_ZoneMotionControl", Zone := "ZoneCounterGbl", Carrier := 11, SDCOUT_DriveFwdCmd => "TC_SDC_Out".Zone["ZoneCounterGbl"].Carrier[11].DriveFwdCMD, SDCOUT_DriveCmdSpeed => "TC_SDC_Out".Zone["ZoneCounterGbl"].Carrier[11].DriveCmdSpeed, SDCOUT_NextStopPos => "TC_SDC_Out".Zone["ZoneCounterGbl"].Carrier[11].NextStopPos, SDCOUT_NextCarrierNum => "TC_SDC_Out".Zone["ZoneCounterGbl"].Carrier[11].NextCarrierNum, SDCOut_AtCmdPos => "TC_SDC_Out".Zone["ZoneCounterGbl"].Carrier[11].AtCmdPos)
      "IDB601_MapSDCOut_Carrier_DB"(ZoneArray := "TC_SDC_Out".Zone, Carrier := 11, Zone := "ZoneCounterGbl", DriveFwdCMD => "EMS".Carrier[11].SDC_OUT.DriveFwdCMD, AtCmdPos => "EMS".Carrier[11].SDC_OUT.AtCmdPos, NextStopPos => "EMS".Carrier[11].SDC_OUT.NextStopPos, DriveCmdSpeed => "EMS".Carrier[11].SDC_OUT.DriveCmdSpeed, Zone_Echo => "EMS".Carrier[11].SDC_OUT.Zone, Pos_Echo => "EMS".Carrier[11].SDC_OUT.CarrierPosition)
   END_RUNG
   // the same network as SCL:
   "IDB609_TCMapSDCOutFB"(TC_ZoneMotion := "DB116_TC_ZoneMotionControl",   // "FB118_TCMapSDCOut"
                          Zone := "ZoneCounterGbl",
                          Carrier := 11,
                          SDCOUT_DriveFwdCmd => "TC_SDC_Out".Zone["ZoneCounterGbl"].Carrier[11].DriveFwdCMD,
                          SDCOUT_DriveCmdSpeed => "TC_SDC_Out".Zone["ZoneCounterGbl"].Carrier[11].DriveCmdSpeed,
                          SDCOUT_NextStopPos => "TC_SDC_Out".Zone["ZoneCounterGbl"].Carrier[11].NextStopPos,
                          SDCOUT_NextCarrierNum => "TC_SDC_Out".Zone["ZoneCounterGbl"].Carrier[11].NextCarrierNum,
                          SDCOut_AtCmdPos => "TC_SDC_Out".Zone["ZoneCounterGbl"].Carrier[11].AtCmdPos,
                          ENO => #_w1);
   IF #_w1 THEN
       "IDB601_MapSDCOut_Carrier_DB"(ZoneArray := "TC_SDC_Out".Zone,   // "FB117_MapSDCOut_Carrier"
                               Carrier := 11,
                               Zone := "ZoneCounterGbl",
                               DriveFwdCMD => "EMS".Carrier[11].SDC_OUT.DriveFwdCMD,
                               AtCmdPos => "EMS".Carrier[11].SDC_OUT.AtCmdPos,
                               NextStopPos => "EMS".Carrier[11].SDC_OUT.NextStopPos,
                               DriveCmdSpeed => "EMS".Carrier[11].SDC_OUT.DriveCmdSpeed,
                               Zone_Echo => "EMS".Carrier[11].SDC_OUT.Zone,
                               Pos_Echo => "EMS".Carrier[11].SDC_OUT.CarrierPosition);
   END_IF;
END_REGION

